(* Logix 5000 project; controller PLC_MCC1300_75F1 vendor 1 type 14 code 166 rev 32.11; software revision 32.04; part 30 of 83 *)
(* tags used below, declared in another part *)
   B3 : DINT[51];
   C5 : COUNTER[51];
   CNV8_RES_CAPID : ALIAS FOR N40[8];
   CNV9_FWD : ALIAS FOR O[21].8;
   I : INT[128];   // Local Input Updates Input Slot 2
   N11 : DINT[500];
   N12 : DINT[500];
   N14 : DINT[500];
   N209 : DINT[100];
   N214_1 : ALIAS FOR N214[1];
   N25 : DINT[110];
   N26 : DINT[150];
   N26_101 : ALIAS FOR N26[101];
   N7 : DINT[101];
   O : INT[128];
   QC3_PE : ALIAS FOR B3[6].12;
   QC3_PE_N : ALIAS FOR B3[13].0;
   T4 : TIMER[51];
   TMP_d : DINT;
   VIN_A_INSP_S1 : ALIAS FOR N26[30].0;
   VIN_GRP_ID : ALIAS FOR N26[0];
   VIN_LEN_S1 : ALIAS FOR N26[21];
   VIN_NTOL_WID : ALIAS FOR N26[11];
   VIN_NUM_SPLITS : ALIAS FOR N26[4];
   VIN_NUM_STRMS : ALIAS FOR N26[3];
   VIN_PTOL_WID : ALIAS FOR N26[5];
   VIN_SUB_THICK : ALIAS FOR N26[2];
   VIN_SUB_TYPE : ALIAS FOR N26[1];
   VIN_WID_A : ALIAS FOR N26[17];
   VIS_IGNORE_LEN_EN : ALIAS FOR N26[100].12;
   VIS_OUTPT_OFF : ALIAS FOR N27[60].2;
   VIS_SYS_STOPPED : ALIAS FOR N27[60].1;
   VOUT_GRP_ID : ALIAS FOR N27[0];
   VOUT_NEW_DATA : ALIAS FOR N27[2];
   VRES_GRP_ID : ALIAS FOR N25[0];
   VRES_REJ_1A : ALIAS FOR N25[5];
   xAlwaysOFF : BOOL;
(* MainProgram, continued *)

ROUTINE _4_VIS_INTFCE   (* ladder *)
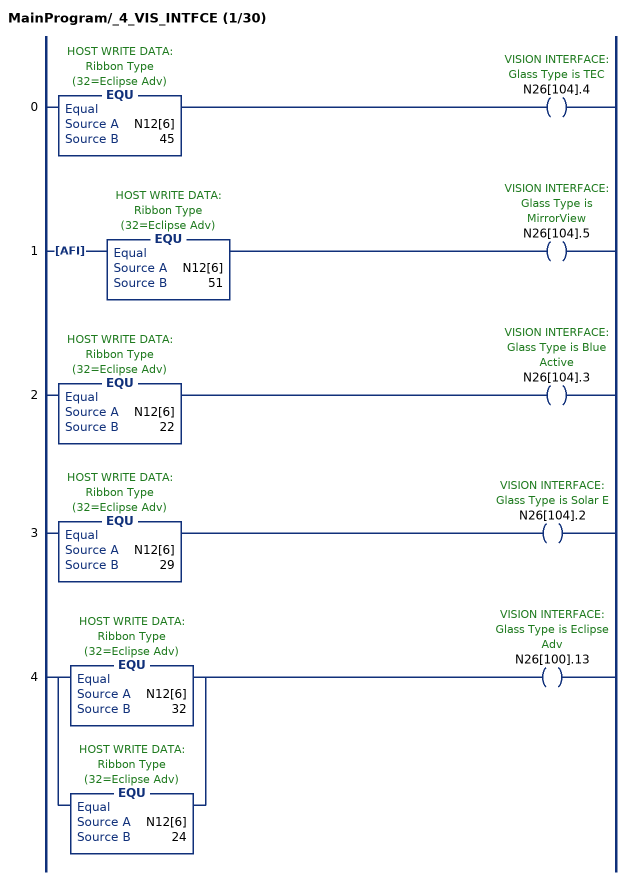
   0: EQU(N12[6],45)OTE(N26[104].4);
   1: AFI()EQU(N12[6],51)OTE(N26[104].5);
   2: EQU(N12[6],22)OTE(N26[104].3);
   3: EQU(N12[6],29)OTE(N26[104].2);
   4: [EQU(N12[6],32) ,EQU(N12[6],24) ]OTE(N26[100].13);
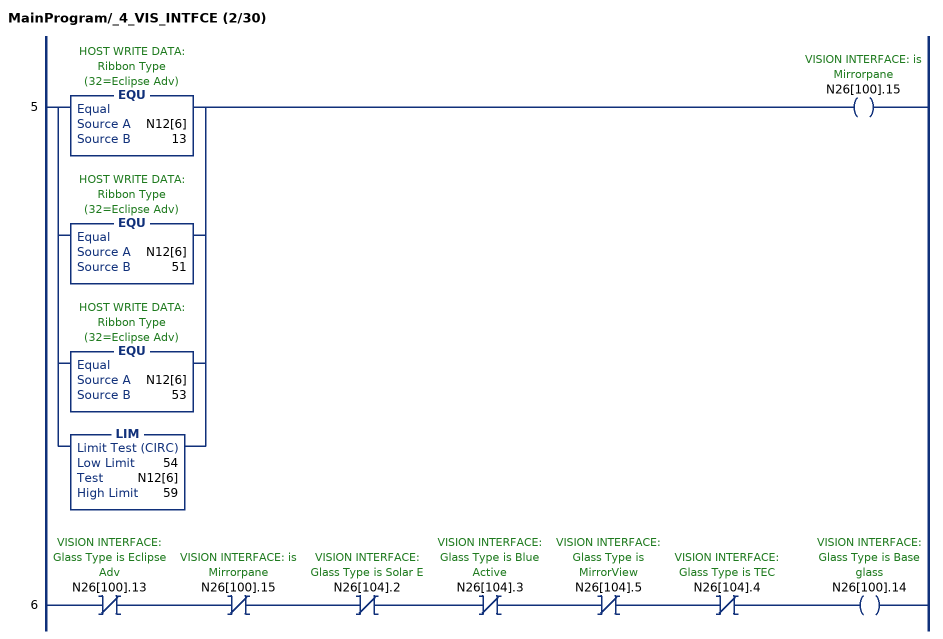
   5: [EQU(N12[6],13) ,EQU(N12[6],51) ,EQU(N12[6],53) ,LIM(54,N12[6],59) ]OTE(N26[100].15);
   6: XIO(N26[100].13)XIO(N26[100].15)XIO(N26[104].2)XIO(N26[104].3)XIO(N26[104].5)XIO(N26[104].4)OTE(N26[100].14);
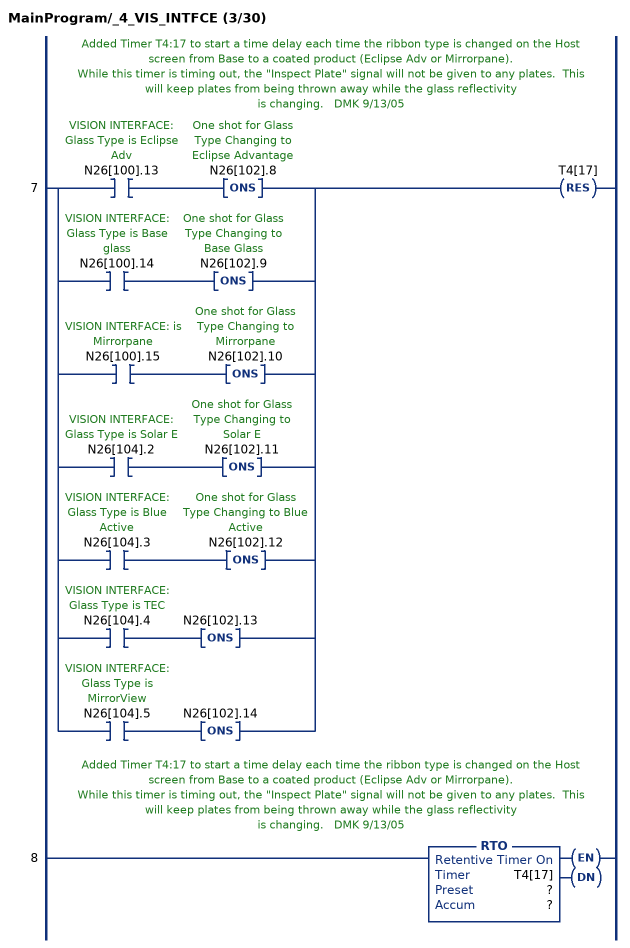
   // Added Timer T4:17 to start a time delay each time the ribbon type is changed on the Host screen from Base to a coated product (Eclipse Adv or Mirrorpane).
   // While this timer is timing out, the "Inspect Plate" signal will not be given to any plates.  This will keep plates from being thrown away while the glass reflectivity
   // is changing.   DMK 9/13/05
   7: [XIC(N26[100].13) ONS(N26[102].8) ,XIC(N26[100].14) ONS(N26[102].9) ,XIC(N26[100].15) ONS(N26[102].10) ,XIC(N26[104].2) ONS(N26[102].11) ,XIC(N26[104].3) ONS(N26[102].12) ,XIC(N26[104].4) ONS(N26[102].13) ,XIC(N26[104].5) ONS(N26[102].14) ]RES(T4[17]);
   // Added Timer T4:17 to start a time delay each time the ribbon type is changed on the Host screen from Base to a coated product (Eclipse Adv or Mirrorpane).
   // While this timer is timing out, the "Inspect Plate" signal will not be given to any plates.  This will keep plates from being thrown away while the glass reflectivity
   // is changing.   DMK 9/13/05
   8: RTO(T4[17],?,?);
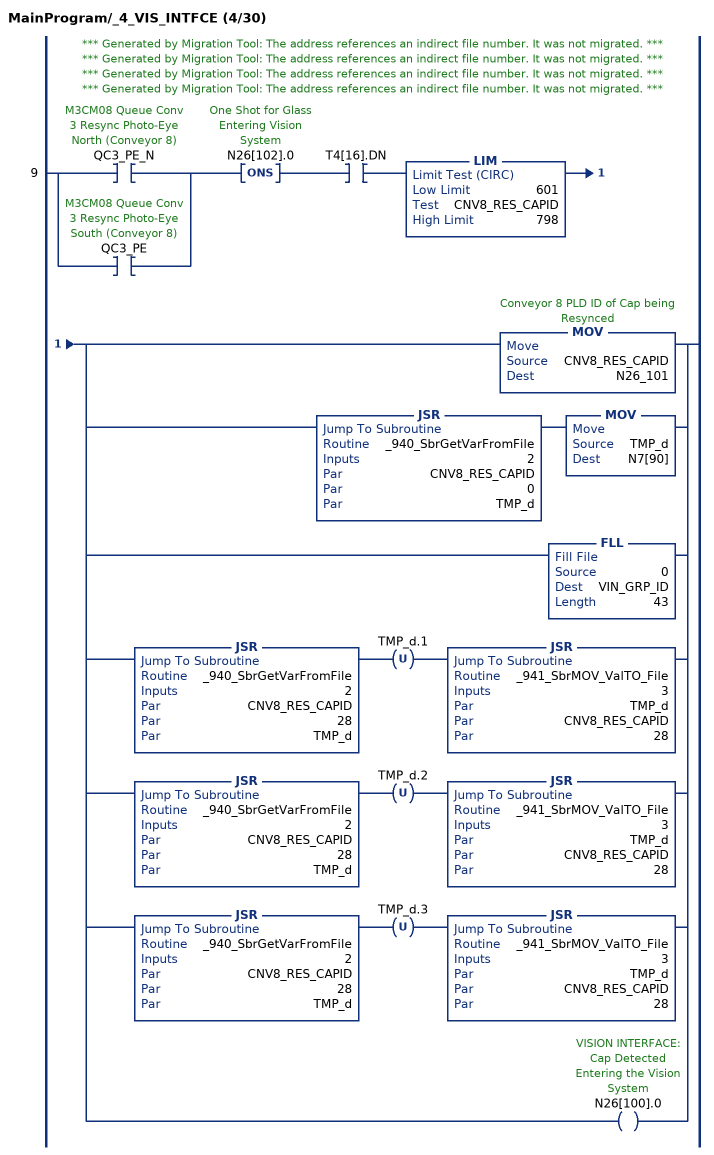
   // *** Generated by Migration Tool: The address references an indirect file number. It was not migrated. ***
   // *** Generated by Migration Tool: The address references an indirect file number. It was not migrated. ***
   // *** Generated by Migration Tool: The address references an indirect file number. It was not migrated. ***
   // *** Generated by Migration Tool: The address references an indirect file number. It was not migrated. ***
   9: [XIC(QC3_PE_N) ,XIC(QC3_PE) ]ONS(N26[102].0)XIC(T4[16].DN)LIM(601,CNV8_RES_CAPID,798)[MOV(CNV8_RES_CAPID,N26_101) ,JSR(_940_SbrGetVarFromFile,2,CNV8_RES_CAPID,0,TMP_d) MOV(TMP_d,N7[90]) ,FLL(0,VIN_GRP_ID,43) ,JSR(_940_SbrGetVarFromFile,2,CNV8_RES_CAPID,28,TMP_d) OTU(TMP_d.1) JSR(_941_SbrMOV_ValTO_File,3,TMP_d,CNV8_RES_CAPID,28) ,JSR(_940_SbrGetVarFromFile,2,CNV8_RES_CAPID,28,TMP_d) OTU(TMP_d.2) JSR(_941_SbrMOV_ValTO_File,3,TMP_d,CNV8_RES_CAPID,28) ,JSR(_940_SbrGetVarFromFile,2,CNV8_RES_CAPID,28,TMP_d) OTU(TMP_d.3) JSR(_941_SbrMOV_ValTO_File,3,TMP_d,CNV8_RES_CAPID,28) ,OTE(N26[100].0) ];
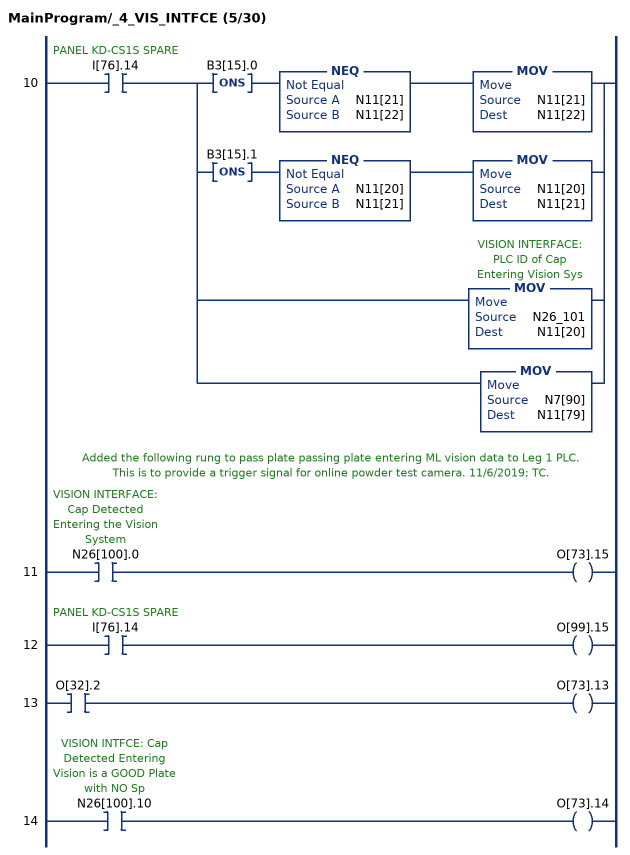
   10: XIC(I[76].14)[ONS(B3[15].0) NEQ(N11[21],N11[22]) MOV(N11[21],N11[22]) ,ONS(B3[15].1) NEQ(N11[20],N11[21]) MOV(N11[20],N11[21]) ,MOV(N26_101,N11[20]) ,MOV(N7[90],N11[79]) ];
   // Added the following rung to pass plate passing plate entering ML vision data to Leg 1 PLC. This is to provide a trigger signal for online powder test camera. 11/6/2019; TC.
   11: XIC(N26[100].0)OTE(O[73].15);
   12: XIC(I[76].14)OTE(O[99].15);
   13: XIC(O[32].2)OTE(O[73].13);
   14: XIC(N26[100].10)OTE(O[73].14);
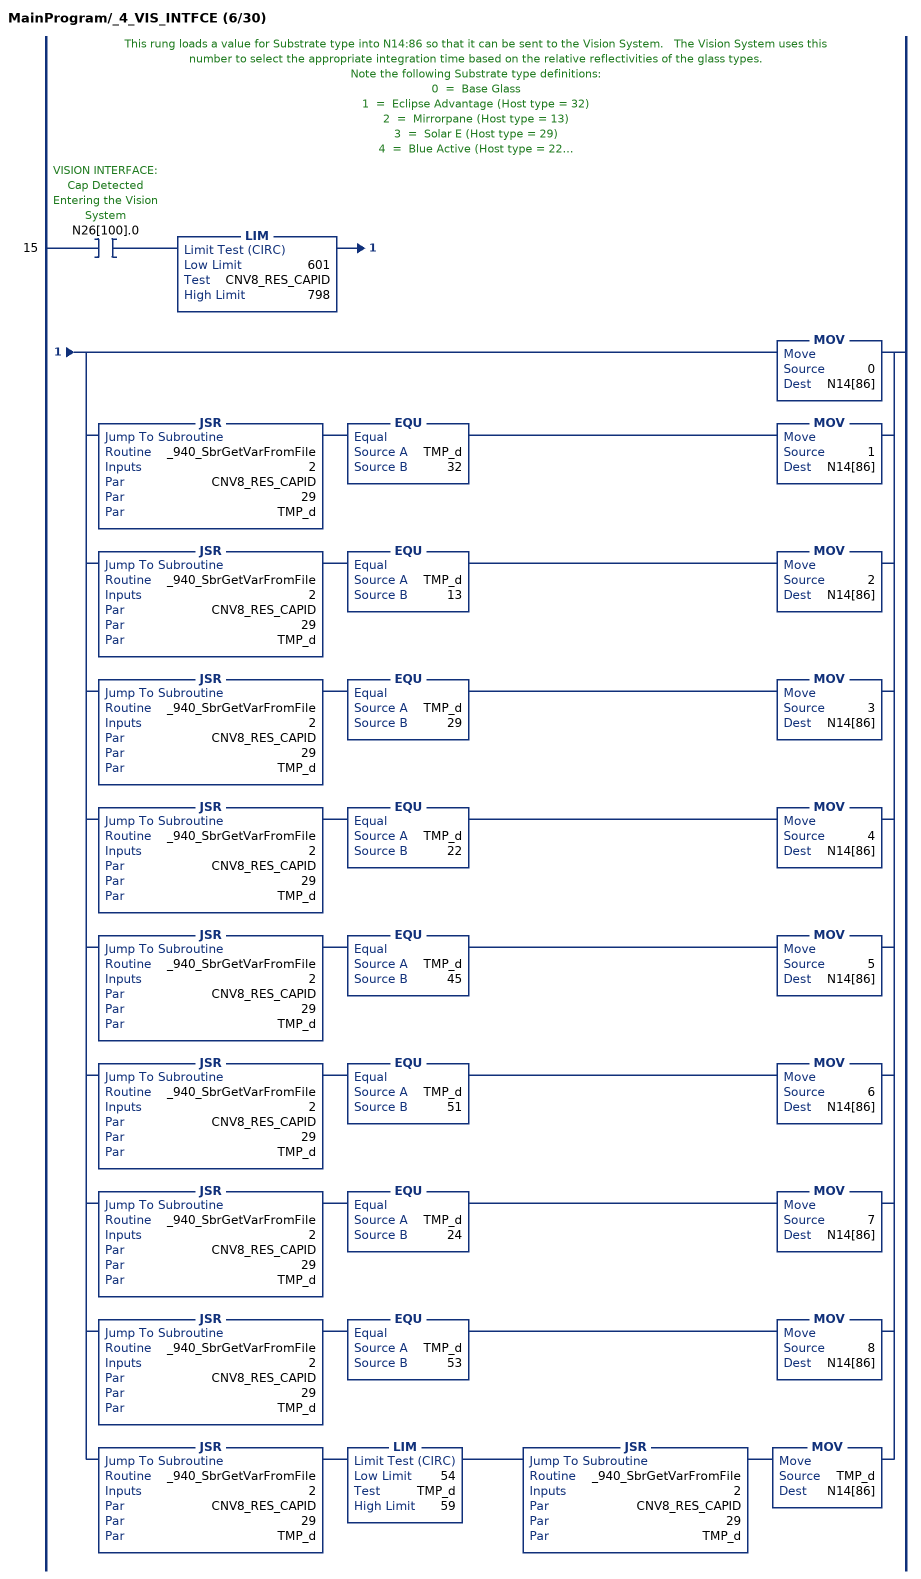
   // This rung loads a value for Substrate type into N14:86 so that it can be sent to the Vision System.   The Vision System uses this
   // number to select the appropriate integration time based on the relative reflectivities of the glass types.
   // Note the following Substrate type definitions:
   //  0  =  Base Glass
   //  1  =  Eclipse Advantage (Host type = 32)
   //  2  =  Mirrorpane (Host type = 13)
   //  3  =  Solar E (Host type = 29)
   //  4  =  Blue Active (Host type = 22)
   // *** Generated by Migration Tool: The address references an indirect file number. It was not migrated. ***
   // *** Generated by Migration Tool: The address references an indirect file number. It was not migrated. ***
   // *** Generated by Migration Tool: The address references an indirect file number. It was not migrated. ***
   // *** Generated by Migration Tool: The address references an indirect file number. It was not migrated. ***
   // *** Generated by Migration Tool: The address references an indirect file number. It was not migrated. ***
   // *** Generated by Migration Tool: The address references an indirect file number. It was not migrated. ***
   // *** Generated by Migration Tool: The address references an indirect file number. It was not migrated. ***
   // *** Generated by Migration Tool: The address references an indirect file number. It was not migrated. ***
   // *** Generated by Migration Tool: The address references an indirect file number. It was not migrated. ***
   // *** Generated by Migration Tool: The address references an indirect file number. It was not migrated. ***
   15: XIC(N26[100].0)LIM(601,CNV8_RES_CAPID,798)[MOV(0,N14[86]) ,JSR(_940_SbrGetVarFromFile,2,CNV8_RES_CAPID,29,TMP_d) EQU(TMP_d,32) MOV(1,N14[86]) ,JSR(_940_SbrGetVarFromFile,2,CNV8_RES_CAPID,29,TMP_d) EQU(TMP_d,13) MOV(2,N14[86]) ,JSR(_940_SbrGetVarFromFile,2,CNV8_RES_CAPID,29,TMP_d) EQU(TMP_d,29) MOV(3,N14[86]) ,JSR(_940_SbrGetVarFromFile,2,CNV8_RES_CAPID,29,TMP_d) EQU(TMP_d,22) MOV(4,N14[86]) ,JSR(_940_SbrGetVarFromFile,2,CNV8_RES_CAPID,29,TMP_d) EQU(TMP_d,45) MOV(5,N14[86]) ,JSR(_940_SbrGetVarFromFile,2,CNV8_RES_CAPID,29,TMP_d) EQU(TMP_d,51) MOV(6,N14[86]) ,JSR(_940_SbrGetVarFromFile,2,CNV8_RES_CAPID,29,TMP_d) EQU(TMP_d,24) MOV(7,N14[86]) ,JSR(_940_SbrGetVarFromFile,2,CNV8_RES_CAPID,29,TMP_d) EQU(TMP_d,53) MOV(8,N14[86]) ,JSR(_940_SbrGetVarFromFile,2,CNV8_RES_CAPID,29,TMP_d) LIM(54,TMP_d,59) JSR(_940_SbrGetVarFromFile,2,CNV8_RES_CAPID,29,TMP_d) MOV(TMP_d,N14[86]) ];
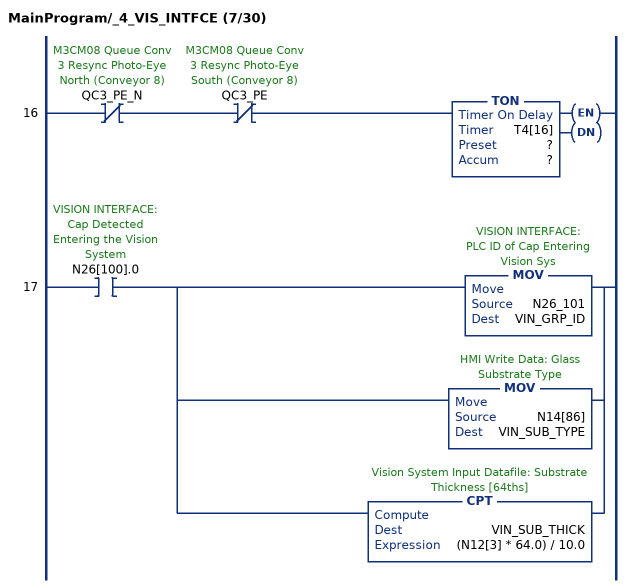
   16: XIO(QC3_PE_N)XIO(QC3_PE)TON(T4[16],?,?);
   17: XIC(N26[100].0)[MOV(N26_101,VIN_GRP_ID) ,MOV(N14[86],VIN_SUB_TYPE) ,CPT(VIN_SUB_THICK,(N12[3] * 64.0) / 10.0) ];
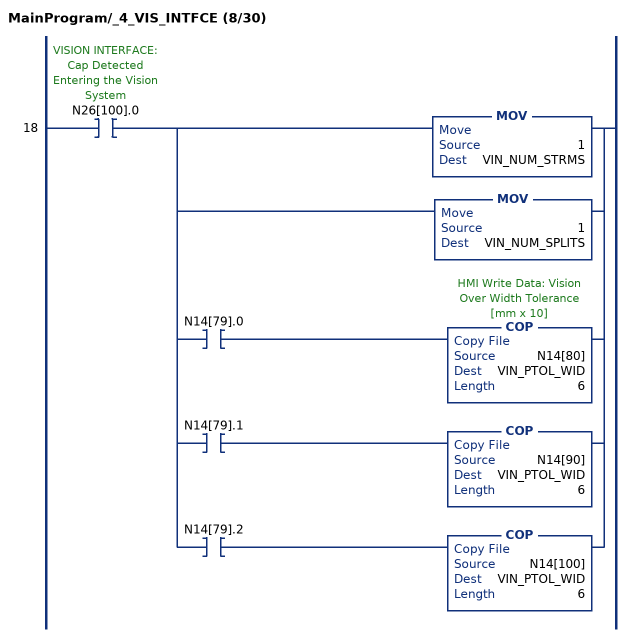
   18: XIC(N26[100].0)[MOV(1,VIN_NUM_STRMS) ,MOV(1,VIN_NUM_SPLITS) ,XIC(N14[79].0) COP(N14[80],VIN_PTOL_WID,6) ,XIC(N14[79].1) COP(N14[90],VIN_PTOL_WID,6) ,XIC(N14[79].2) COP(N14[100],VIN_PTOL_WID,6) ];
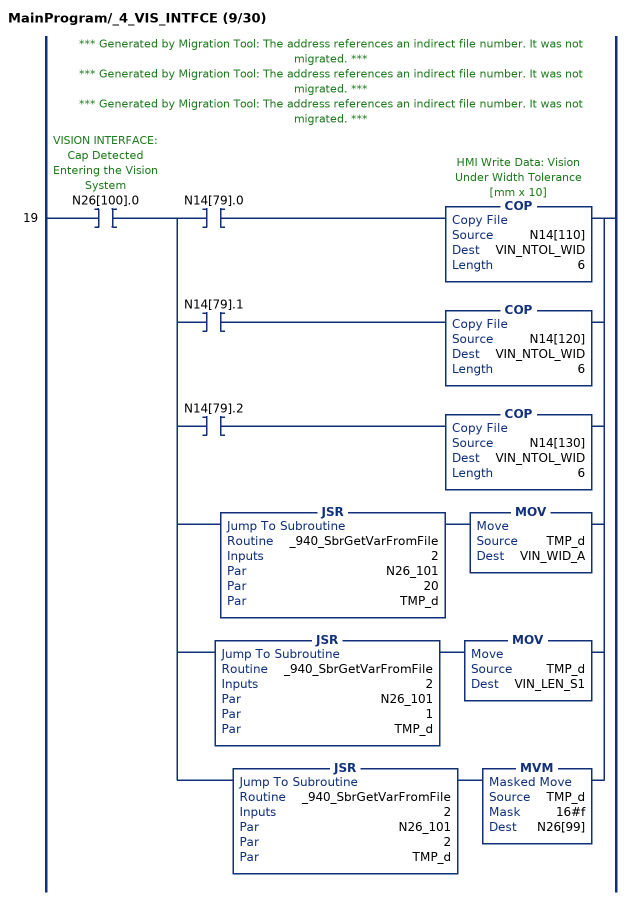
   // *** Generated by Migration Tool: The address references an indirect file number. It was not migrated. ***
   // *** Generated by Migration Tool: The address references an indirect file number. It was not migrated. ***
   // *** Generated by Migration Tool: The address references an indirect file number. It was not migrated. ***
   19: XIC(N26[100].0)[XIC(N14[79].0) COP(N14[110],VIN_NTOL_WID,6) ,XIC(N14[79].1) COP(N14[120],VIN_NTOL_WID,6) ,XIC(N14[79].2) COP(N14[130],VIN_NTOL_WID,6) ,JSR(_940_SbrGetVarFromFile,2,N26_101,20,TMP_d) MOV(TMP_d,VIN_WID_A) ,JSR(_940_SbrGetVarFromFile,2,N26_101,1,TMP_d) MOV(TMP_d,VIN_LEN_S1) ,JSR(_940_SbrGetVarFromFile,2,N26_101,2,TMP_d) MVM(TMP_d,16#f,N26[99]) ];
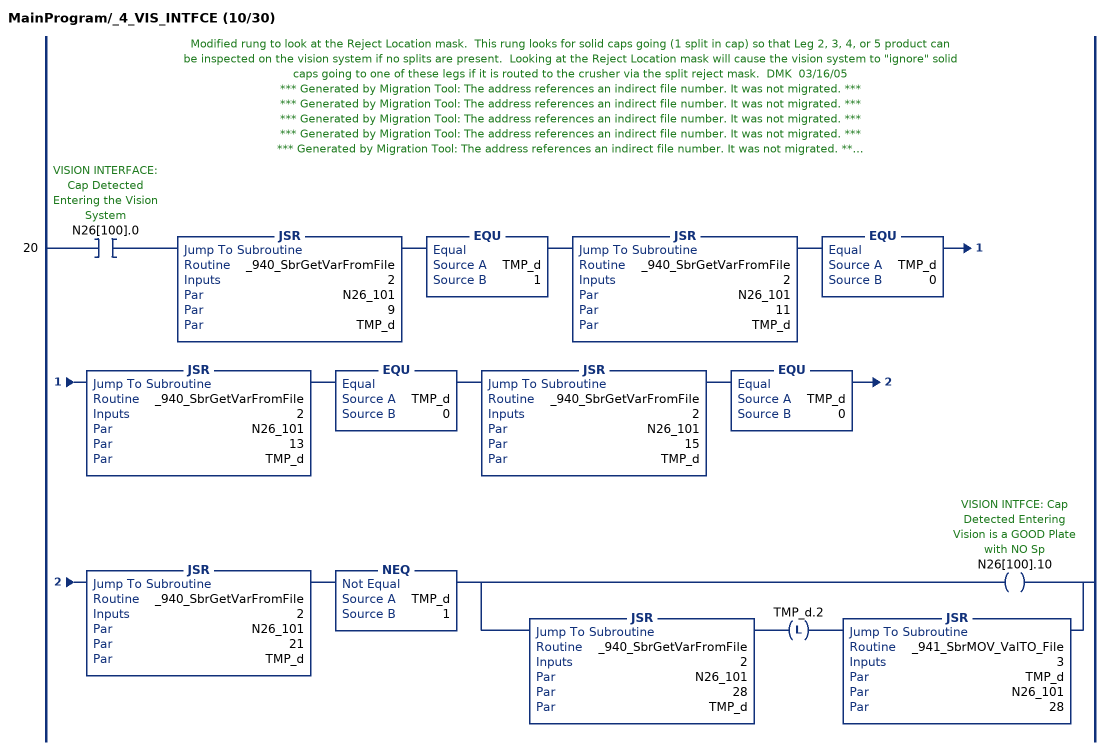
   // Modified rung to look at the Reject Location mask.  This rung looks for solid caps going (1 split in cap) so that Leg 2, 3, 4, or 5 product can
   // be inspected on the vision system if no splits are present.  Looking at the Reject Location mask will cause the vision system to "ignore" solid
   // caps going to one of these legs if it is routed to the crusher via the split reject mask.  DMK  03/16/05
   // *** Generated by Migration Tool: The address references an indirect file number. It was not migrated. ***
   // *** Generated by Migration Tool: The address references an indirect file number. It was not migrated. ***
   // *** Generated by Migration Tool: The address references an indirect file number. It was not migrated. ***
   // *** Generated by Migration Tool: The address references an indirect file number. It was not migrated. ***
   // *** Generated by Migration Tool: The address references an indirect file number. It was not migrated. ***
   // *** Generated by Migration Tool: The address references an indirect file number. It was not migrated. ***
   20: XIC(N26[100].0)JSR(_940_SbrGetVarFromFile,2,N26_101,9,TMP_d)EQU(TMP_d,1)JSR(_940_SbrGetVarFromFile,2,N26_101,11,TMP_d)EQU(TMP_d,0)JSR(_940_SbrGetVarFromFile,2,N26_101,13,TMP_d)EQU(TMP_d,0)JSR(_940_SbrGetVarFromFile,2,N26_101,15,TMP_d)EQU(TMP_d,0)JSR(_940_SbrGetVarFromFile,2,N26_101,21,TMP_d)NEQ(TMP_d,1)[OTE(N26[100].10) ,JSR(_940_SbrGetVarFromFile,2,N26_101,28,TMP_d) OTL(TMP_d.2) JSR(_941_SbrMOV_ValTO_File,3,TMP_d,N26_101,28) ];
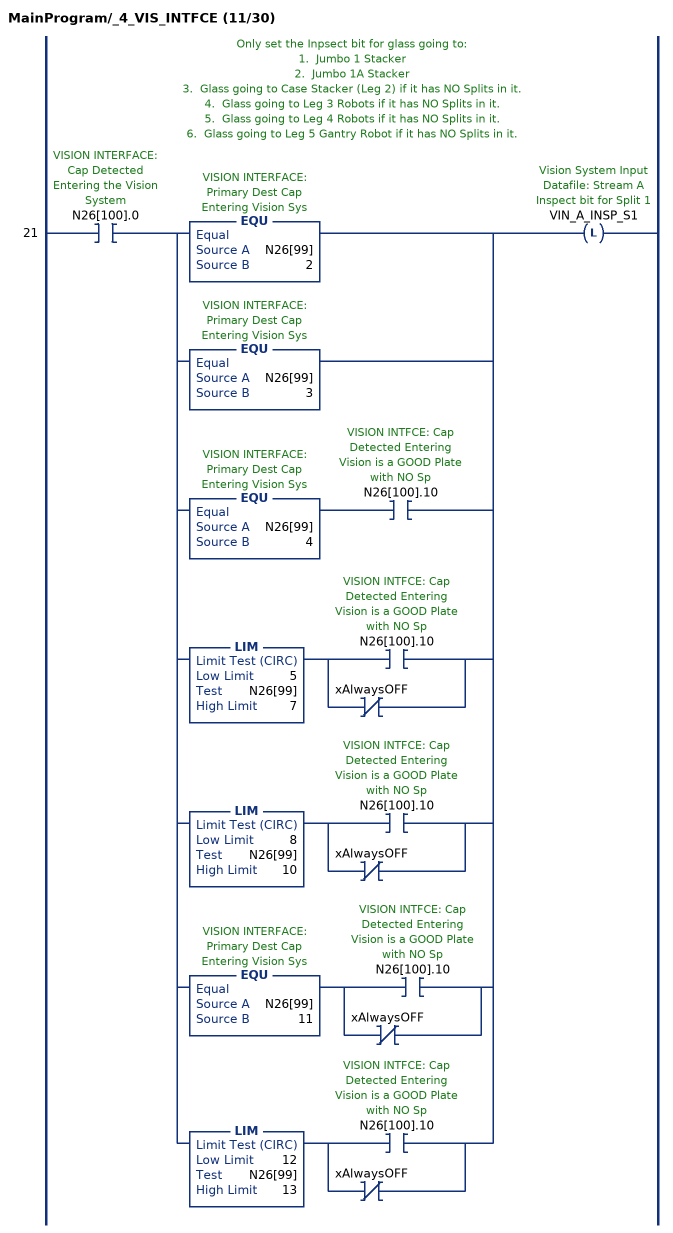
   // Only set the Inpsect bit for glass going to:
   // 1.  Jumbo 1 Stacker
   // 2.  Jumbo 1A Stacker
   // 3.  Glass going to Case Stacker (Leg 2) if it has NO Splits in it.
   // 4.  Glass going to Leg 3 Robots if it has NO Splits in it.
   // 5.  Glass going to Leg 4 Robots if it has NO Splits in it.
   // 6.  Glass going to Leg 5 Gantry Robot if it has NO Splits in it.
   21: XIC(N26[100].0)[EQU(N26[99],2) ,EQU(N26[99],3) ,EQU(N26[99],4) XIC(N26[100].10) ,LIM(5,N26[99],7) [XIC(N26[100].10) ,XIO(xAlwaysOFF) ] ,LIM(8,N26[99],10) [XIC(N26[100].10) ,XIO(xAlwaysOFF) ] ,EQU(N26[99],11) [XIC(N26[100].10) ,XIO(xAlwaysOFF) ] ,LIM(12,N26[99],13) [XIC(N26[100].10) ,XIO(xAlwaysOFF) ] ]OTL(VIN_A_INSP_S1);
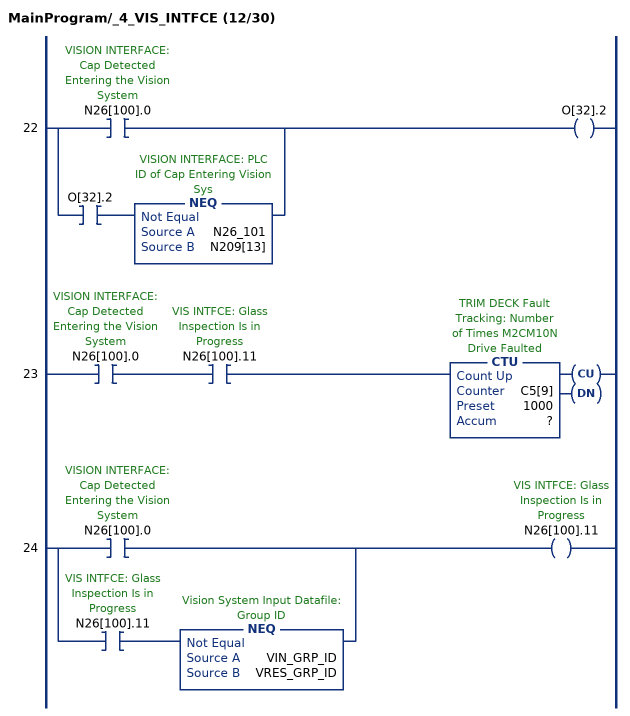
   22: [XIC(N26[100].0) ,XIC(O[32].2) NEQ(N26_101,N209[13]) ]OTE(O[32].2);
   23: XIC(N26[100].0)XIC(N26[100].11)CTU(C5[9],?,?);
   24: [XIC(N26[100].0) ,XIC(N26[100].11) NEQ(VIN_GRP_ID,VRES_GRP_ID) ]OTE(N26[100].11);
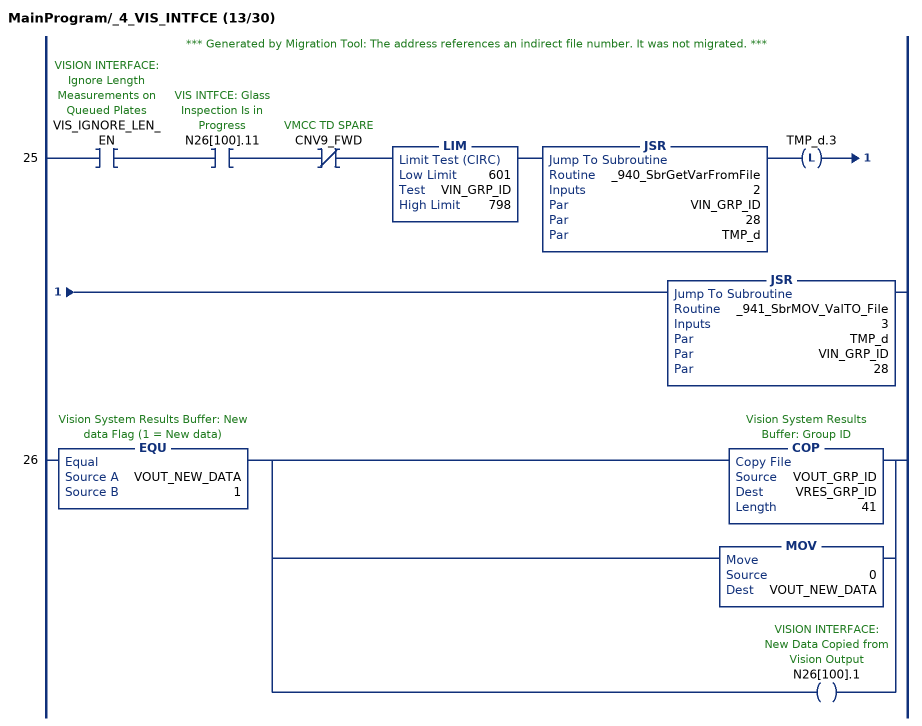
   // *** Generated by Migration Tool: The address references an indirect file number. It was not migrated. ***
   25: XIC(VIS_IGNORE_LEN_EN)XIC(N26[100].11)XIO(CNV9_FWD)LIM(601,VIN_GRP_ID,798)JSR(_940_SbrGetVarFromFile,2,VIN_GRP_ID,28,TMP_d)OTL(TMP_d.3)JSR(_941_SbrMOV_ValTO_File,3,TMP_d,VIN_GRP_ID,28);
   26: EQU(VOUT_NEW_DATA,1)[COP(VOUT_GRP_ID,VRES_GRP_ID,41) ,MOV(0,VOUT_NEW_DATA) ,OTE(N26[100].1) ];
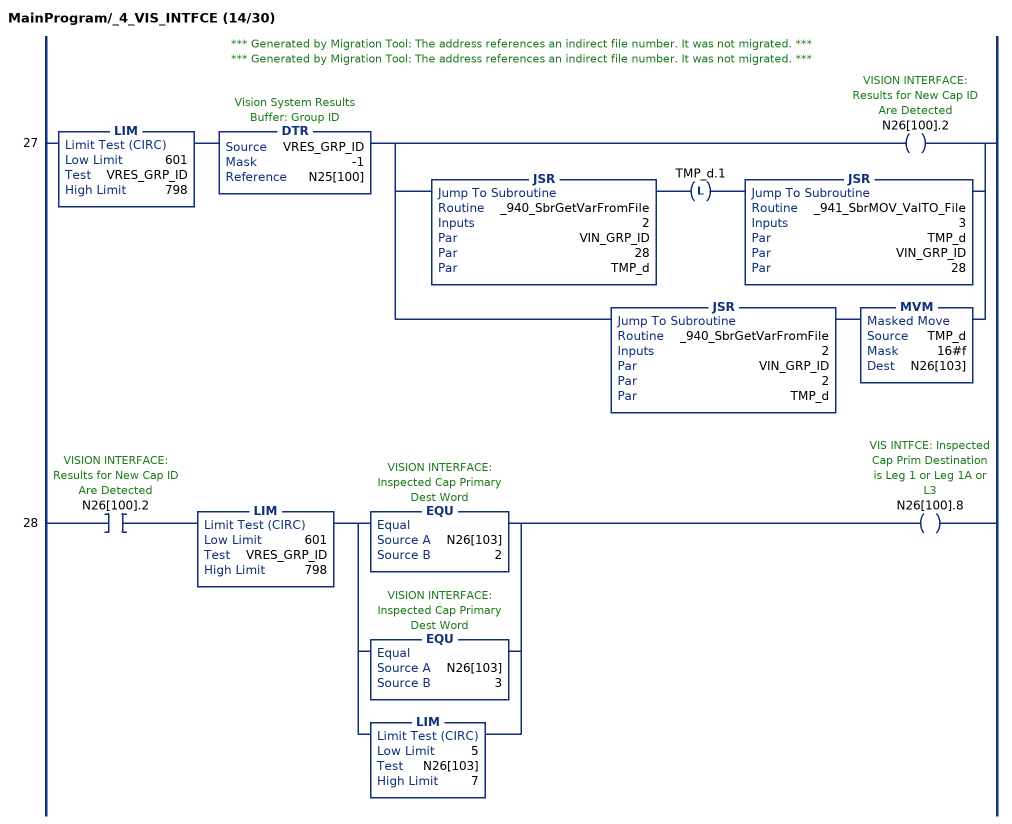
   // *** Generated by Migration Tool: The address references an indirect file number. It was not migrated. ***
   // *** Generated by Migration Tool: The address references an indirect file number. It was not migrated. ***
   27: LIM(601,VRES_GRP_ID,798)DTR(VRES_GRP_ID,-1,N25[100])[OTE(N26[100].2) ,JSR(_940_SbrGetVarFromFile,2,VIN_GRP_ID,28,TMP_d) OTL(TMP_d.1) JSR(_941_SbrMOV_ValTO_File,3,TMP_d,VIN_GRP_ID,28) ,JSR(_940_SbrGetVarFromFile,2,VIN_GRP_ID,2,TMP_d) MVM(TMP_d,16#f,N26[103]) ];
   28: XIC(N26[100].2)LIM(601,VRES_GRP_ID,798)[EQU(N26[103],2) ,EQU(N26[103],3) ,LIM(5,N26[103],7) ]OTE(N26[100].8);